   TextField "Text field_22" at 649,435 size 53x20; Text 'IW230'
   Button "HmiScreenItemData_8" at 469,45 size 355x40; TextOn 'Back'; TextOff 'Text'
   TextField "Screen title" at 455,41 size 373x50; Text 'Screen title'

screen "RIO 4 Analogue Settings" 1280x800, template "Template"
   on GenerateScreen: "TitleUpdater"()
   Button "HmiScreenItemData_1" at 1,1 size 150x40; TextOn 'Back'; TextOff 'Commissioning'
      on Release: ActivateScreen("Commissioning Main Page", 0)
   TextField "Text field_82" at 60,138 size 215x20; Text 'Tank 4P USD Flow FIT-418-4P'
   TextField "Text field_90" at 286,114 size 62x18; Text 'Reading'
   IOField "I/O field_2" at 281,138 size 75x20; FormatPattern 999; Unit  Nm³/hr
      ProcessValue <- "20_TANKS_IP_DATA_RIO_04_FIRST_TANK_USD_FLOW"
   TextField "Text field_1" at 359,114 size 68x18; Text 'Low Low'
   TextField "Text field_2" at 442,114 size 34x18; Text 'Low'
   TextField "Text field_3" at 509,114 size 37x18; Text 'High'
   TextField "Text field_4" at 561,114 size 74x18; Text 'High High'
   TextField "Text field_5" at 434,92 size 74x18; Text 'Setpoints'
   TextField "Text field_6" at 7,138 size 53x20; Text 'IW260'
   TextField "Text field_7" at 60,175 size 215x20; Text 'Tank 4P MBG Flow FIT-420-4P'
   IOField "I/O field_6" at 281,175 size 75x20; FormatPattern 999; Unit  Nm³/hr
      ProcessValue <- "20_TANKS_IP_DATA_RIO_04_FIRST_TANK_MBG_FLOW"
   TextField "Text field_8" at 7,175 size 53x20; Text 'IW262'
   TextField "Text field_9" at 60,212 size 215x20; Text 'Tank 4S USD Flow FIT-417-4S'
   IOField "I/O field_11" at 281,212 size 75x20; FormatPattern 999; Unit  Nm³/hr
      ProcessValue <- "20_TANKS_IP_DATA_RIO_04_SECOND_TANK_USD_FLOW"
   TextField "Text field_10" at 7,212 size 53x20; Text 'IW264'
   TextField "Text field_11" at 60,249 size 215x20; Text 'Tank 4S MBG Flow FIT-419-4S'
   IOField "I/O field_16" at 281,249 size 75x20; FormatPattern 999; Unit  Nm³/hr
      ProcessValue <- "20_TANKS_IP_DATA_RIO_04_SECOND_TANK_MBG_FLOW"
   TextField "Text field_12" at 7,249 size 53x20; Text 'IW266'
   TextField "Text field_13" at 60,286 size 215x20; Text 'RIO 4 Deck Main Pressure PT-415'
   TextField "Text field_14" at 7,286 size 53x20; Text 'IW268'
   TextField "Text field_15" at 60,324 size 215x20; Text 'Tank 4P BW Level LT-422-4P'
   TextField "Text field_16" at 7,324 size 53x20; Text 'IW270'
   TextField "Text field_17" at 60,361 size 215x20; Text 'Tank 4S BW Level LT-421-4S'
   TextField "Text field_18" at 7,361 size 53x20; Text 'IW272'
   TextField "Text field_25" at 702,324 size 215x20; Text 'Tank 4S BW Temperature 425-4S'
   TextField "Text field_26" at 928,114 size 62x18; Text 'Reading'
   IOField "I/O field_51" at 922,324 size 75x20; FormatPattern s999.9; Unit  °C
      ProcessValue <- "20_TANKS_IP_DATA_RIO_04_SECOND_TANK_BWT_TEMP"
   TextField "Text field_27" at 1001,114 size 68x18; Text 'Low Low'
   TextField "Text field_28" at 1082,114 size 34x18; Text 'Low'
   TextField "Text field_29" at 1150,114 size 37x18; Text 'High'
   TextField "Text field_30" at 1203,114 size 74x18; Text 'High High'
   TextField "Text field_31" at 1076,92 size 74x18; Text 'Setpoints'
   TextField "Text field_32" at 649,324 size 53x20; Text 'IW286'
   TextField "Text field_33" at 702,361 size 215x20; Text 'Tank 4S BW DO TX-427-4S'
   IOField "I/O field_56" at 922,361 size 75x20; FormatPattern 99.9; Unit  mg/l
      ProcessValue <- "20_TANKS_IP_DATA_RIO_04_SECOND_TANK_BWT_DO"
   TextField "Text field_34" at 649,361 size 53x20; Text 'IW288'
   TextField "Text field_35" at 702,398 size 215x20; Text 'Confined Space O2 Level Port'
   IOField "I/O field_61" at 922,398 size 75x20; FormatPattern 99.9; Unit  %
      ProcessValue <- "20_TANKS_IP_DATA_RIO_04_FIRST_TANK_O2_MONITOR"
   TextField "Text field_36" at 649,398 size 53x20; Text 'IW290'
   TextField "Text field_65" at 702,138 size 215x20; Text 'Tank 4P BW ph TX-426-4P'
   IOField "I/O field_126" at 922,138 size 75x20; FormatPattern 999.9
      ProcessValue <- "20_TANKS_IP_DATA_RIO_04_FIRST_TANK_BWT_PH"
   TextField "Text field_66" at 649,138 size 53x20; Text 'IW276'
   TextField "Text field_67" at 702,175 size 215x20; Text 'Tank 4P BW Temperature 426-4P'
   IOField "I/O field_131" at 922,175 size 75x20; FormatPattern s999.9; Unit  °C
      ProcessValue <- "20_TANKS_IP_DATA_RIO_04_FIRST_TANK_BWT_TEMP"
   TextField "Text field_68" at 649,175 size 53x20; Text 'IW278'
   TextField "Text field_69" at 702,212 size 215x20; Text 'Tank 4P BW DO TX-428-4P'
   IOField "I/O field_136" at 922,212 size 75x20; FormatPattern 99.9; Unit  mg/l
      ProcessValue <- "20_TANKS_IP_DATA_RIO_04_FIRST_TANK_BWT_DO"
   TextField "Text field_70" at 649,212 size 53x20; Text 'IW280'
   TextField "Text field_71" at 702,249 size 215x20; Text 'RIO 4 Tanks Pressure PT-424'
   TextField "Text field_72" at 649,249 size 53x20; Text 'IW282'
   TextField "Text field_73" at 702,286 size 215x20; Text 'Tank 4S BW ph TX-425-4S'
   IOField "I/O field_146" at 922,286 size 75x20; FormatPattern 999.9
      ProcessValue <- "20_TANKS_IP_DATA_RIO_04_SECOND_TANK_BWT_PH"
   TextField "Text field_74" at 649,286 size 53x20; Text 'IW284'
   TextField "Text field_41" at 133,114 size 85x18; Text 'Description'
   TextField "Text field_42" at 771,114 size 85x18; Text 'Description'
   TextField "Text field_43" at 17,114 size 21x18; Text 'AI'
   TextField "Text field_44" at 661,114 size 21x18; Text 'AI'
   IOField "I/O field_21" at 281,285 size 75x20; FormatPattern 99.9; Unit  Bar
      ProcessValue <- "20_TANKS_IP_DATA_RIO_04_FIRST_TANK_DECK_IG_PRESS"
   IOField "I/O field_26" at 281,322 size 75x20; FormatPattern 999.9; Unit  %
      ProcessValue <- "20_TANKS_IP_DATA_RIO_04_FIRST_TANK_BWT_LEVEL"
   IOField "I/O field_27" at 281,359 size 75x20; FormatPattern 999.9; Unit  %
      ProcessValue <- "20_TANKS_IP_DATA_RIO_04_SECOND_TANK_BWT_LEVEL"
   IOField "I/O field_93" at 922,249 size 75x20; FormatPattern s999.9; Unit  mBar
      ProcessValue <- "20_TANKS_IP_DATA_RIO_04_FIRST_TANK_TANKS_PRESS"
   TextField "Text field_21" at 702,435 size 215x20; Text 'Confined Space O2 Level Starboard'
   IOField "I/O field_41" at 922,435 size 75x20; FormatPattern 99.9; Unit  %
      ProcessValue <- "20_TANKS_IP_DATA_RIO_04_SECOND_TANK_O2_MONITOR"
   TextField "Text field_22" at 649,435 size 53x20; Text 'IW290'
   IOField "I/O field_1" at 361,138 size 60x20; Authorization "User administration"; FormatPattern 999
      ProcessValue <- "2084_Setpoints_FIT418_LoLo"
   IOField "I/O field_3" at 429,138 size 60x20; Authorization "User administration"; FormatPattern 999
      ProcessValue <- "2084_Setpoints_FIT418_Lo"
   IOField "I/O field_4" at 497,138 size 60x20; Authorization "User administration"; FormatPattern 999
      ProcessValue <- "2084_Setpoints_FIT418_Hi"
   IOField "I/O field_5" at 565,138 size 60x20; Authorization "User administration"; FormatPattern 999
      ProcessValue <- "2084_Setpoints_FIT418_HiHi"
   IOField "I/O field_7" at 361,175 size 60x20; FormatPattern 999
      ProcessValue <- "2084_Setpoints_FIT420_LoLo"
   IOField "I/O field_8" at 429,175 size 60x20; FormatPattern 999
      ProcessValue <- "2084_Setpoints_FIT420_Lo"
   IOField "I/O field_9" at 497,175 size 60x20; Authorization "User administration"; FormatPattern 999
      ProcessValue <- "2084_Setpoints_FIT420_Hi"
   IOField "I/O field_10" at 565,175 size 60x20; Authorization "User administration"; FormatPattern 999
      ProcessValue <- "2084_Setpoints_FIT420_HiHi"
   IOField "I/O field_12" at 361,212 size 60x20; FormatPattern 999
      ProcessValue <- "2084_Setpoints_FIT417_LoLo"
   IOField "I/O field_13" at 429,212 size 60x20; FormatPattern 999
      ProcessValue <- "2084_Setpoints_FIT417_Lo"
   IOField "I/O field_14" at 497,212 size 60x20; Authorization "User administration"; FormatPattern 999
      ProcessValue <- "2084_Setpoints_FIT417_Hi"
   IOField "I/O field_15" at 565,212 size 60x20; Authorization "User administration"; FormatPattern 999
      ProcessValue <- "2084_Setpoints_FIT417_HiHi"
   IOField "I/O field_17" at 361,249 size 60x20; FormatPattern 999
      ProcessValue <- "2084_Setpoints_FIT419_LoLo"
   IOField "I/O field_18" at 429,249 size 60x20; FormatPattern 999
      ProcessValue <- "2084_Setpoints_FIT419_Lo"
   IOField "I/O field_19" at 497,249 size 60x20; FormatPattern 999
      ProcessValue <- "2084_Setpoints_FIT419_Hi"
   IOField "I/O field_20" at 565,249 size 60x20; FormatPattern 999
      ProcessValue <- "2084_Setpoints_FIT419_HiHi"
   IOField "I/O field_22" at 361,285 size 60x20; FormatPattern 99.999
      ProcessValue <- "2084_Setpoints_PIT415_LoLo"
   IOField "I/O field_23" at 429,285 size 60x20; FormatPattern 99.999
      ProcessValue <- "2084_Setpoints_PIT415_Lo"
   IOField "I/O field_24" at 497,285 size 60x20; FormatPattern 99.999
      ProcessValue <- "2084_Setpoints_PIT415_Hi"
   IOField "I/O field_25" at 565,285 size 60x20; FormatPattern 99.999
      ProcessValue <- "2084_Setpoints_PIT415_HiHi"
   IOField "I/O field_28" at 429,359 size 60x20; Authorization "User administration"; FormatPattern 999
      ProcessValue <- "2084_Setpoints_LT421_Lo"
   IOField "I/O field_29" at 497,359 size 60x20; Authorization "User administration"; FormatPattern 999
      ProcessValue <- "2084_Setpoints_LT421_Hi"
   IOField "I/O field_30" at 429,322 size 60x20; Authorization "User administration"; FormatPattern 999
      ProcessValue <- "2084_Setpoints_LT422_Lo"
   IOField "I/O field_31" at 497,322 size 60x20; Authorization "User administration"; FormatPattern 999
      ProcessValue <- "2084_Setpoints_LT422_Hi"
   IOField "I/O field_32" at 361,322 size 60x20; FormatPattern 9.9
   IOField "I/O field_33" at 361,359 size 60x20; FormatPattern 9.9
   IOField "I/O field_34" at 565,322 size 60x20; FormatPattern 9.9
   IOField "I/O field_35" at 565,359 size 60x20; FormatPattern 9.9
   IOField "I/O field_62" at 1004,397 size 60x20; FormatPattern 99.9
      ProcessValue <- "2084_Setpoints_Conf O2 Level Lo Lo"
   IOField "I/O field_63" at 1072,397 size 60x20; FormatPattern 99.9
      ProcessValue <- "2084_Setpoints_Conf O2 Level Lo"
   IOField "I/O field_64" at 1139,397 size 60x20; Authorization "User administration"; FormatPattern 99.9
   IOField "I/O field_65" at 1207,397 size 60x20; Authorization "User administration"; FormatPattern 99.9
   IOField "I/O field_72" at 1004,286 size 60x20; FormatPattern 99.9
   IOField "I/O field_74" at 1004,323 size 60x20; FormatPattern 99.9
   IOField "I/O field_75" at 1072,323 size 60x20; FormatPattern 99.9
   IOField "I/O field_77" at 1207,286 size 60x20; Authorization "User administration"; FormatPattern 99.9
   IOField "I/O field_78" at 1139,323 size 60x20; Authorization "User administration"; FormatPattern 99.9
   IOField "I/O field_79" at 1207,323 size 60x20; Authorization "User administration"; FormatPattern 99.9
   IOField "I/O field_80" at 1139,360 size 60x20; Authorization "User administration"; FormatPattern 99.9
      ProcessValue <- "2084_Setpoints_TX427 Star DO High"
   IOField "I/O field_86" at 1207,360 size 60x20; Authorization "User administration"; FormatPattern 99.9
   IOField "I/O field_87" at 1004,360 size 60x20; Authorization "User administration"; FormatPattern 99.9
   IOField "I/O field_88" at 1072,360 size 60x20; Authorization "User administration"; FormatPattern 99.9
      ProcessValue <- "2084_Setpoints_TX427 Star DO Lo"
   IOField "I/O field_52" at 1003,138 size 60x20; FormatPattern 99.9
   IOField "I/O field_53" at 1071,138 size 60x20; FormatPattern 99.9
      ProcessValue <- "2084_Setpoints_TX426 Port PH Lo"
   IOField "I/O field_54" at 1003,175 size 60x20; FormatPattern 99.9
   IOField "I/O field_55" at 1071,175 size 60x20; FormatPattern 99.9
   IOField "I/O field_57" at 1139,138 size 60x20; Authorization "User administration"; FormatPattern 99.9
      ProcessValue <- "2084_Setpoints_TX426 Port PH High"
   IOField "I/O field_58" at 1207,138 size 60x20; Authorization "User administration"; FormatPattern 99.9
   IOField "I/O field_59" at 1139,175 size 60x20; Authorization "User administration"; FormatPattern 99.9
   IOField "I/O field_60" at 1207,175 size 60x20; Authorization "User administration"; FormatPattern 99.9
   IOField "I/O field_89" at 1139,212 size 60x20; Authorization "User administration"; FormatPattern 99.9
      ProcessValue <- "2084_Setpoints_TX428 Port DO High"
   IOField "I/O field_90" at 1207,212 size 60x20; Authorization "User administration"; FormatPattern 99.9
   IOField "I/O field_91" at 1003,212 size 60x20; Authorization "User administration"; FormatPattern 99.9
   IOField "I/O field_92" at 1071,212 size 60x20; Authorization "User administration"; FormatPattern 99.9
      ProcessValue <- "2084_Setpoints_TX428 Port DO Lo"
   IOField "I/O field_94" at 1139,249 size 60x20; Authorization "User administration"; FormatPattern 999.9
      ProcessValue <- "2084_Setpoints_PIT424_Hi"
   IOField "I/O field_95" at 1207,249 size 60x20; Authorization "User administration"; FormatPattern 999.9
      ProcessValue <- "2084_Setpoints_PIT424_HiHi"
   IOField "I/O field_96" at 1004,249 size 60x20; Authorization "User administration"; FormatPattern 999.9
      ProcessValue <- "2084_Setpoints_PIT424_LoLo"
   IOField "I/O field_97" at 1072,249 size 60x20; Authorization "User administration"; FormatPattern 999.9
      ProcessValue <- "2084_Setpoints_PIT424_Lo"
   IOField "I/O field_42" at 1072,286 size 60x20; FormatPattern 99.9
      ProcessValue <- "2084_Setpoints_TX425 Star PH Lo"
   IOField "I/O field_43" at 1139,286 size 60x20; Authorization "User administration"; FormatPattern 99.9
      ProcessValue <- "2084_Setpoints_TX425 Star PH High"
   Group "Group" at 455,41 size 373x50
   Button "HmiScreenItemData_8" at 469,45 size 355x40; TextOn 'Back'; TextOff 'Text'
   TextField "Screen title" at 455,41 size 373x50; Text 'Screen title'

screen "RIO 5 Analogue Settings" 1280x800, template "Template"
   on GenerateScreen: "TitleUpdater"()
   Button "HmiScreenItemData_1" at 1,1 size 150x40; TextOn 'Back'; TextOff 'Commissioning'
      on Release: ActivateScreen("Commissioning Main Page", 0)
   TextField "Text field_82" at 60,138 size 215x20; Text 'Tank 5P USD Flow FIT-418-5P'
   TextField "Text field_90" at 286,114 size 62x18; Text 'Reading'
   IOField "I/O field_2" at 281,138 size 75x20; FormatPattern 999; Unit  Nm³/hr
      ProcessValue <- "20_TANKS_IP_DATA_RIO_05_FIRST_TANK_USD_FLOW"
   TextField "Text field_1" at 359,114 size 68x18; Text 'Low Low'
   TextField "Text field_2" at 442,114 size 34x18; Text 'Low'
   TextField "Text field_3" at 509,114 size 37x18; Text 'High'
   TextField "Text field_4" at 561,114 size 74x18; Text 'High High'
   TextField "Text field_5" at 434,92 size 74x18; Text 'Setpoints'
   TextField "Text field_6" at 7,138 size 53x20; Text 'IW300'
   TextField "Text field_7" at 60,175 size 215x20; Text 'Tank 5P MBG Flow FIT-420-5P'
   IOField "I/O field_6" at 281,175 size 75x20; FormatPattern 999; Unit  Nm³/hr
      ProcessValue <- "20_TANKS_IP_DATA_RIO_05_FIRST_TANK_MBG_FLOW"
   TextField "Text field_8" at 7,175 size 53x20; Text 'IW302'
   TextField "Text field_9" at 60,212 size 215x20; Text 'Tank 5S USD Flow FIT-417-5S'
   IOField "I/O field_11" at 281,212 size 75x20; FormatPattern 999; Unit  Nm³/hr
      ProcessValue <- "20_TANKS_IP_DATA_RIO_05_SECOND_TANK_USD_FLOW"
   TextField "Text field_10" at 7,212 size 53x20; Text 'IW304'
   TextField "Text field_11" at 60,249 size 215x20; Text 'Tank 5S MBG Flow FIT-419-5S'
   IOField "I/O field_16" at 281,249 size 75x20; FormatPattern 999; Unit  Nm³/hr
      ProcessValue <- "20_TANKS_IP_DATA_RIO_05_SECOND_TANK_MBG_FLOW"
   TextField "Text field_12" at 7,249 size 53x20; Text 'IW306'
   TextField "Text field_13" at 60,286 size 215x20; Text 'RIO 5 Deck Main Pressure PT-415'
   TextField "Text field_14" at 7,286 size 53x20; Text 'IW308'
   TextField "Text field_15" at 60,324 size 215x20; Text 'Tank 5P BW Level LT-422-5P'
   TextField "Text field_16" at 7,324 size 53x20; Text 'IW310'
   TextField "Text field_17" at 60,361 size 215x20; Text 'Tank 5S BW Level LT-421-5S'
   TextField "Text field_18" at 7,361 size 53x20; Text 'IW312'
   TextField "Text field_25" at 702,324 size 215x20; Text 'Tank 5S BW Temperature 425-5S'
   TextField "Text field_26" at 928,114 size 62x18; Text 'Reading'
   IOField "I/O field_51" at 922,324 size 75x20; FormatPattern s999.9; Unit  °C
      ProcessValue <- "20_TANKS_IP_DATA_RIO_05_SECOND_TANK_BWT_TEMP"
   TextField "Text field_27" at 1001,114 size 68x18; Text 'Low Low'
   TextField "Text field_28" at 1082,114 size 34x18; Text 'Low'
   TextField "Text field_29" at 1150,114 size 37x18; Text 'High'
   TextField "Text field_30" at 1203,114 size 74x18; Text 'High High'
   TextField "Text field_31" at 1076,92 size 74x18; Text 'Setpoints'
   TextField "Text field_32" at 649,324 size 53x20; Text 'IW326'
   TextField "Text field_33" at 702,361 size 215x20; Text 'Tank 5S BW DO TX-427-5S'
   IOField "I/O field_56" at 922,361 size 75x20; FormatPattern 99.9; Unit  mg/l
      ProcessValue <- "20_TANKS_IP_DATA_RIO_05_SECOND_TANK_BWT_DO"
   TextField "Text field_34" at 649,361 size 53x20; Text 'IW328'
   TextField "Text field_35" at 702,398 size 215x20; Text 'Confined Space Oxygen Level'
   IOField "I/O field_61" at 922,398 size 75x20; FormatPattern 99.9; Unit  %
      ProcessValue <- "20_TANKS_IP_DATA_RIO_05_FIRST_TANK_O2_MONITOR"
   TextField "Text field_36" at 649,398 size 53x20; Text 'IW330'
   TextField "Text field_65" at 702,138 size 215x20; Text 'Tank 5P BW ph TX-426-5P'
   IOField "I/O field_126" at 922,138 size 75x20; FormatPattern 99.9
      ProcessValue <- "20_TANKS_IP_DATA_RIO_05_FIRST_TANK_BWT_PH"
   TextField "Text field_66" at 649,138 size 53x20; Text 'IW316'
   TextField "Text field_67" at 702,175 size 215x20; Text 'Tank 5P BW Temperature 426-5P'
   IOField "I/O field_131" at 922,175 size 75x20; FormatPattern s999.9; Unit  °C
      ProcessValue <- "20_TANKS_IP_DATA_RIO_05_FIRST_TANK_BWT_TEMP"
   TextField "Text field_68" at 649,175 size 53x20; Text 'IW318'
   TextField "Text field_69" at 702,212 size 215x20; Text 'Tank 5P BW DO TX-428-5P'
   IOField "I/O field_136" at 922,212 size 75x20; FormatPattern s99.99; Unit  mg/l
      ProcessValue <- "20_TANKS_IP_DATA_RIO_05_FIRST_TANK_BWT_DO"
   TextField "Text field_70" at 649,212 size 53x20; Text 'IW320'
   TextField "Text field_71" at 702,249 size 215x20; Text 'RIO 5 Tanks Pressure PT-424'
   TextField "Text field_72" at 649,249 size 53x20; Text 'IW322'
   TextField "Text field_73" at 702,286 size 215x20; Text 'Tank 5S BW ph TX-425-5S'
   IOField "I/O field_146" at 922,286 size 75x20; FormatPattern 99.9
      ProcessValue <- "20_TANKS_IP_DATA_RIO_05_SECOND_TANK_BWT_PH"
   TextField "Text field_74" at 649,286 size 53x20; Text 'IW324'
   TextField "Text field_41" at 133,114 size 85x18; Text 'Description'
   TextField "Text field_42" at 771,114 size 85x18; Text 'Description'
   TextField "Text field_43" at 17,114 size 21x18; Text 'AI'
   TextField "Text field_44" at 661,114 size 21x18; Text 'AI'
   IOField "I/O field_21" at 281,285 size 75x20; FormatPattern 99.999; Unit  Bar
      ProcessValue <- "20_TANKS_IP_DATA_RIO_05_FIRST_TANK_DECK_IG_PRESS"
   IOField "I/O field_26" at 281,322 size 75x20; FormatPattern 999.9; Unit  %
      ProcessValue <- "20_TANKS_IP_DATA_RIO_05_FIRST_TANK_BWT_LEVEL"
   IOField "I/O field_27" at 281,359 size 75x20; FormatPattern 999.9; Unit  %
      ProcessValue <- "20_TANKS_IP_DATA_RIO_05_SECOND_TANK_BWT_LEVEL"
   IOField "I/O field_93" at 922,249 size 75x20; FormatPattern 999.9; Unit  mBar
      ProcessValue <- "20_TANKS_IP_DATA_RIO_05_FIRST_TANK_TANKS_PRESS"
   Group "Group" at 455,41 size 373x50
   TextField "Text field_21" at 702,435 size 215x20; Text 'Confined Space Oxygen Level'
   IOField "I/O field_41" at 922,435 size 75x20; FormatPattern 99.9; Unit  %
      ProcessValue <- "20_TANKS_IP_DATA_RIO_05_SECOND_TANK_O2_MONITOR"
   TextField "Text field_22" at 649,435 size 53x20; Text 'IW330'
   IOField "I/O field_1" at 361,138 size 60x20; Authorization "User administration"; FormatPattern 999
      ProcessValue <- "2084_Setpoints_FIT418_LoLo"
   IOField "I/O field_3" at 429,138 size 60x20; Authorization "User administration"; FormatPattern 999
      ProcessValue <- "2084_Setpoints_FIT418_Lo"
   IOField "I/O field_4" at 497,138 size 60x20; Authorization "User administration"; FormatPattern 999
      ProcessValue <- "2084_Setpoints_FIT418_Hi"
   IOField "I/O field_5" at 565,138 size 60x20; Authorization "User administration"; FormatPattern 999
      ProcessValue <- "2084_Setpoints_FIT418_HiHi"
   IOField "I/O field_7" at 361,175 size 60x20; FormatPattern 999
      ProcessValue <- "2084_Setpoints_FIT420_LoLo"
   IOField "I/O field_8" at 429,175 size 60x20; FormatPattern 999
      ProcessValue <- "2084_Setpoints_FIT420_Lo"
   IOField "I/O field_9" at 497,175 size 60x20; Authorization "User administration"; FormatPattern 999
      ProcessValue <- "2084_Setpoints_FIT420_Hi"
   IOField "I/O field_10" at 565,175 size 60x20; Authorization "User administration"; FormatPattern 999
      ProcessValue <- "2084_Setpoints_FIT420_HiHi"
   IOField "I/O field_12" at 361,212 size 60x20; FormatPattern 999
      ProcessValue <- "2084_Setpoints_FIT417_LoLo"
   IOField "I/O field_13" at 429,212 size 60x20; FormatPattern 999
      ProcessValue <- "2084_Setpoints_FIT417_Lo"
   IOField "I/O field_14" at 497,212 size 60x20; Authorization "User administration"; FormatPattern 999
      ProcessValue <- "2084_Setpoints_FIT417_Hi"
   IOField "I/O field_15" at 565,212 size 60x20; Authorization "User administration"; FormatPattern 999
      ProcessValue <- "2084_Setpoints_FIT417_HiHi"
   IOField "I/O field_17" at 361,249 size 60x20; FormatPattern 999
      ProcessValue <- "2084_Setpoints_FIT419_LoLo"
   IOField "I/O field_18" at 429,249 size 60x20; FormatPattern 999
      ProcessValue <- "2084_Setpoints_FIT419_Lo"
   IOField "I/O field_19" at 497,249 size 60x20; FormatPattern 999
      ProcessValue <- "2084_Setpoints_FIT419_Hi"
   IOField "I/O field_20" at 565,249 size 60x20; FormatPattern 999
      ProcessValue <- "2084_Setpoints_FIT419_HiHi"
   IOField "I/O field_22" at 361,285 size 60x20; FormatPattern 99.999
      ProcessValue <- "2084_Setpoints_PIT415_LoLo"
   IOField "I/O field_23" at 429,285 size 60x20; FormatPattern 99.999
      ProcessValue <- "2084_Setpoints_PIT415_Lo"
   IOField "I/O field_24" at 497,285 size 60x20; FormatPattern 99.999
      ProcessValue <- "2084_Setpoints_PIT415_Hi"
   IOField "I/O field_25" at 565,285 size 60x20; FormatPattern 99.999
      ProcessValue <- "2084_Setpoints_PIT415_HiHi"
   IOField "I/O field_28" at 429,359 size 60x20; Authorization "User administration"; FormatPattern 999
      ProcessValue <- "2084_Setpoints_LT421_Lo"
   IOField "I/O field_29" at 497,359 size 60x20; Authorization "User administration"; FormatPattern 999
      ProcessValue <- "2084_Setpoints_LT421_Hi"
   IOField "I/O field_30" at 429,322 size 60x20; Authorization "User administration"; FormatPattern 999
      ProcessValue <- "2084_Setpoints_LT422_Lo"
   IOField "I/O field_31" at 497,322 size 60x20; Authorization "User administration"; FormatPattern 999
      ProcessValue <- "2084_Setpoints_LT422_Hi"
   IOField "I/O field_32" at 361,322 size 60x20; FormatPattern 9.9
   IOField "I/O field_33" at 361,359 size 60x20; FormatPattern 9.9
   IOField "I/O field_34" at 565,322 size 60x20; FormatPattern 9.9
   IOField "I/O field_35" at 565,359 size 60x20; FormatPattern 9.9
   IOField "I/O field_62" at 1004,397 size 60x20; FormatPattern 99.9
      ProcessValue <- "2084_Setpoints_Conf O2 Level Lo Lo"
   IOField "I/O field_63" at 1072,397 size 60x20; FormatPattern 99.9
      ProcessValue <- "2084_Setpoints_Conf O2 Level Lo"
   IOField "I/O field_64" at 1139,397 size 60x20; Authorization "User administration"; FormatPattern 99.9
   IOField "I/O field_65" at 1207,397 size 60x20; Authorization "User administration"; FormatPattern 99.9
   IOField "I/O field_72" at 1004,286 size 60x20; FormatPattern 99.9
   IOField "I/O field_74" at 1004,323 size 60x20; FormatPattern 99.9
   IOField "I/O field_75" at 1072,323 size 60x20; FormatPattern 99.9
   IOField "I/O field_77" at 1207,286 size 60x20; Authorization "User administration"; FormatPattern 99.9
   IOField "I/O field_78" at 1139,323 size 60x20; Authorization "User administration"; FormatPattern 99.9
   IOField "I/O field_79" at 1207,323 size 60x20; Authorization "User administration"; FormatPattern 99.9
   IOField "I/O field_80" at 1139,360 size 60x20; Authorization "User administration"; FormatPattern 99.9
      ProcessValue <- "2084_Setpoints_TX427 Star DO High"
   IOField "I/O field_86" at 1207,360 size 60x20; Authorization "User administration"; FormatPattern 99.9
   IOField "I/O field_87" at 1004,360 size 60x20; Authorization "User administration"; FormatPattern 99.9
   IOField "I/O field_88" at 1072,360 size 60x20; Authorization "User administration"; FormatPattern 99.9
      ProcessValue <- "2084_Setpoints_TX427 Star DO Lo"
   IOField "I/O field_52" at 1003,138 size 60x20; FormatPattern 99.9
   IOField "I/O field_53" at 1071,138 size 60x20; FormatPattern 99.9
      ProcessValue <- "2084_Setpoints_TX426 Port PH Lo"
   IOField "I/O field_54" at 1003,175 size 60x20; FormatPattern 99.9
   IOField "I/O field_55" at 1071,175 size 60x20; FormatPattern 99.9
   IOField "I/O field_57" at 1139,138 size 60x20; Authorization "User administration"; FormatPattern 99.9
      ProcessValue <- "2084_Setpoints_TX426 Port PH High"
   IOField "I/O field_58" at 1207,138 size 60x20; Authorization "User administration"; FormatPattern 99.9
   IOField "I/O field_59" at 1139,175 size 60x20; Authorization "User administration"; FormatPattern 99.9
   IOField "I/O field_60" at 1207,175 size 60x20; Authorization "User administration"; FormatPattern 99.9
   IOField "I/O field_89" at 1139,212 size 60x20; Authorization "User administration"; FormatPattern 99.9
      ProcessValue <- "2084_Setpoints_TX428 Port DO High"
   IOField "I/O field_90" at 1207,212 size 60x20; Authorization "User administration"; FormatPattern 99.9
   IOField "I/O field_91" at 1003,212 size 60x20; Authorization "User administration"; FormatPattern 99.9
   IOField "I/O field_92" at 1071,212 size 60x20; Authorization "User administration"; FormatPattern 99.9
      ProcessValue <- "2084_Setpoints_TX428 Port DO Lo"
   IOField "I/O field_94" at 1139,249 size 60x20; Authorization "User administration"; FormatPattern 999.9
      ProcessValue <- "2084_Setpoints_PIT424_Hi"
   IOField "I/O field_95" at 1207,249 size 60x20; Authorization "User administration"; FormatPattern 999.9
      ProcessValue <- "2084_Setpoints_PIT424_HiHi"
   IOField "I/O field_96" at 1004,249 size 60x20; Authorization "User administration"; FormatPattern 999.9
      ProcessValue <- "2084_Setpoints_PIT424_LoLo"
   IOField "I/O field_97" at 1072,249 size 60x20; Authorization "User administration"; FormatPattern 999.9
      ProcessValue <- "2084_Setpoints_PIT424_Lo"
   IOField "I/O field_36" at 1072,286 size 60x20; FormatPattern 99.9
      ProcessValue <- "2084_Setpoints_TX425 Star PH Lo"
   IOField "I/O field_42" at 1139,286 size 60x20; Authorization "User administration"; FormatPattern 99.9
      ProcessValue <- "2084_Setpoints_TX425 Star PH High"
   Button "HmiScreenItemData_8" at 469,45 size 355x40; TextOn 'Back'; TextOff 'Text'
   TextField "Screen title" at 455,41 size 373x50; Text 'Screen title'

screen "RIO 6 Analogue Settings" 1280x800, template "Template"
   on GenerateScreen: "TitleUpdater"()
   Button "HmiScreenItemData_1" at 1,1 size 150x40; TextOn 'Back'; TextOff 'Commissioning'
      on Release: ActivateScreen("Commissioning Main Page", 0)
   TextField "Text field_82" at 60,138 size 215x20; Text 'Tank 6P USD Flow FIT-418-6P'
   TextField "Text field_90" at 286,114 size 62x18; Text 'Reading'
   IOField "I/O field_2" at 281,138 size 75x20; FormatPattern 999; Unit  Nm³/hr
      ProcessValue <- "20_TANKS_IP_DATA_RIO_06_FIRST_TANK_USD_FLOW"
   TextField "Text field_1" at 359,114 size 68x18; Text 'Low Low'
   TextField "Text field_2" at 442,114 size 34x18; Text 'Low'
   TextField "Text field_3" at 509,114 size 37x18; Text 'High'
   TextField "Text field_4" at 561,114 size 74x18; Text 'High High'
   TextField "Text field_5" at 434,92 size 74x18; Text 'Setpoints'
   TextField "Text field_6" at 7,138 size 53x20; Text 'IW360'
   TextField "Text field_7" at 60,175 size 215x20; Text 'Tank 6P MBG Flow FIT-420-6P'
   IOField "I/O field_6" at 281,175 size 75x20; FormatPattern 999; Unit  Nm³/hr
      ProcessValue <- "20_TANKS_IP_DATA_RIO_06_FIRST_TANK_MBG_FLOW"
   TextField "Text field_8" at 7,175 size 53x20; Text 'IW362'
   TextField "Text field_9" at 60,212 size 215x20; Text 'Tank 6S USD Flow FIT-417-6S'
   IOField "I/O field_11" at 281,212 size 75x20; FormatPattern 999; Unit  Nm³/hr
      ProcessValue <- "20_TANKS_IP_DATA_RIO_06_SECOND_TANK_USD_FLOW"
   TextField "Text field_10" at 7,212 size 53x20; Text 'IW364'
   TextField "Text field_11" at 60,249 size 215x20; Text 'Tank 6S MBG Flow FIT-419-6S'
   IOField "I/O field_16" at 281,249 size 75x20; FormatPattern 999; Unit  Nm³/hr
      ProcessValue <- "20_TANKS_IP_DATA_RIO_06_SECOND_TANK_MBG_FLOW"
   TextField "Text field_12" at 7,249 size 53x20; Text 'IW366'
   TextField "Text field_13" at 60,286 size 215x20; Text 'RIO 6 Deck Main Pressure PT-415'
   TextField "Text field_14" at 7,286 size 53x20; Text 'IW368'
   TextField "Text field_15" at 60,324 size 215x20; Text 'Tank 6P BW Level LT-422-6P'
   TextField "Text field_16" at 7,324 size 53x20; Text 'IW370'
   TextField "Text field_17" at 60,361 size 215x20; Text 'Tank 6S BW Level LT-421-6S'
   TextField "Text field_18" at 7,361 size 53x20; Text 'IW372'
   TextField "Text field_25" at 702,324 size 215x20; Text 'Tank 6S BW Temperature 425-6S'
   TextField "Text field_26" at 928,114 size 62x18; Text 'Reading'
   IOField "I/O field_51" at 922,324 size 75x20; FormatPattern s999.9; Unit  °C
      ProcessValue <- "20_TANKS_IP_DATA_RIO_06_SECOND_TANK_BWT_TEMP"
   TextField "Text field_27" at 1001,114 size 68x18; Text 'Low Low'
   TextField "Text field_28" at 1082,114 size 34x18; Text 'Low'
   TextField "Text field_29" at 1150,114 size 37x18; Text 'High'
   TextField "Text field_30" at 1203,114 size 74x18; Text 'High High'
   TextField "Text field_31" at 1076,92 size 74x18; Text 'Setpoints'
   TextField "Text field_32" at 649,324 size 53x20; Text 'IW386'
   TextField "Text field_33" at 702,361 size 215x20; Text 'Tank 6S BW DO TX-427-6S'
   IOField "I/O field_56" at 922,361 size 75x20; FormatPattern 99.9; Unit  mg/l
      ProcessValue <- "20_TANKS_IP_DATA_RIO_06_SECOND_TANK_BWT_DO"
   TextField "Text field_34" at 649,361 size 53x20; Text 'IW388'
   TextField "Text field_35" at 702,398 size 215x20; Text 'Confined Space Oxygen Level'
   IOField "I/O field_61" at 922,398 size 75x20; FormatPattern 99.9; Unit  %
      ProcessValue <- "20_TANKS_IP_DATA_RIO_06_FIRST_TANK_O2_MONITOR"
   TextField "Text field_36" at 649,398 size 53x20; Text 'IW390'
   TextField "Text field_65" at 702,138 size 215x20; Text 'Tank 6P BW ph TX-426-6P'
   IOField "I/O field_126" at 922,138 size 75x20; FormatPattern 99.9
      ProcessValue <- "20_TANKS_IP_DATA_RIO_06_FIRST_TANK_BWT_PH"
   TextField "Text field_66" at 649,138 size 53x20; Text 'IW376'
   TextField "Text field_67" at 702,175 size 215x20; Text 'Tank 6P BW Temperature 426-6P'
   IOField "I/O field_131" at 922,175 size 75x20; FormatPattern s999.9; Unit  °C
      ProcessValue <- "20_TANKS_IP_DATA_RIO_06_FIRST_TANK_BWT_TEMP"
   TextField "Text field_68" at 649,175 size 53x20; Text 'IW378'
   TextField "Text field_69" at 702,212 size 215x20; Text 'Tank 6P BW DO TX-428-6P'
   IOField "I/O field_136" at 922,212 size 75x20; FormatPattern 99.9; Unit  mg/l
      ProcessValue <- "20_TANKS_IP_DATA_RIO_06_FIRST_TANK_BWT_DO"
   TextField "Text field_70" at 649,212 size 53x20; Text 'IW380'
   TextField "Text field_71" at 702,249 size 215x20; Text 'RIO 6 Tanks Pressure PT-424'
   TextField "Text field_72" at 649,249 size 53x20; Text 'IW382'
   TextField "Text field_73" at 702,286 size 215x20; Text 'Tank 6S BW ph TX-425-6S'
   IOField "I/O field_146" at 922,286 size 75x20; FormatPattern 99.9
      ProcessValue <- "20_TANKS_IP_DATA_RIO_06_SECOND_TANK_BWT_PH"
   TextField "Text field_74" at 649,286 size 53x20; Text 'IW384'
   TextField "Text field_41" at 133,114 size 85x18; Text 'Description'
   TextField "Text field_42" at 771,114 size 85x18; Text 'Description'
   TextField "Text field_43" at 17,114 size 21x18; Text 'AI'
   TextField "Text field_44" at 661,114 size 21x18; Text 'AI'
   IOField "I/O field_21" at 281,285 size 75x20; FormatPattern s99.999; Unit  Bar
      ProcessValue <- "20_TANKS_IP_DATA_RIO_06_FIRST_TANK_DECK_IG_PRESS"
   IOField "I/O field_26" at 281,322 size 75x20; FormatPattern 999; Unit  %
      ProcessValue <- "20_TANKS_IP_DATA_RIO_06_FIRST_TANK_BWT_LEVEL"
   IOField "I/O field_27" at 281,359 size 75x20; FormatPattern 999; Unit  %
      ProcessValue <- "20_TANKS_IP_DATA_RIO_06_SECOND_TANK_BWT_LEVEL"
   IOField "I/O field_93" at 922,249 size 75x20; FormatPattern s999.9; Unit  mBar
      ProcessValue <- "20_TANKS_IP_DATA_RIO_06_FIRST_TANK_TANKS_PRESS"
   TextField "Text field_19" at 702,434 size 215x20; Text 'Confined Space Oxygen Level'
   IOField "I/O field_36" at 922,434 size 75x20; FormatPattern 99.9; Unit  %
      ProcessValue <- "20_TANKS_IP_DATA_RIO_06_FIRST_TANK_O2_MONITOR"
   TextField "Text field_20" at 649,434 size 53x20; Text 'IW390'
   IOField "I/O field_1" at 361,138 size 60x20; Authorization "User administration"; FormatPattern 999
      ProcessValue <- "2084_Setpoints_FIT418_LoLo"
   IOField "I/O field_3" at 429,138 size 60x20; Authorization "User administration"; FormatPattern 999
      ProcessValue <- "2084_Setpoints_FIT418_Lo"
   IOField "I/O field_4" at 497,138 size 60x20; Authorization "User administration"; FormatPattern 999
      ProcessValue <- "2084_Setpoints_FIT418_Hi"
   IOField "I/O field_5" at 565,138 size 60x20; Authorization "User administration"; FormatPattern 999
      ProcessValue <- "2084_Setpoints_FIT418_HiHi"
   IOField "I/O field_7" at 361,175 size 60x20; FormatPattern 999
      ProcessValue <- "2084_Setpoints_FIT420_LoLo"
   IOField "I/O field_8" at 429,175 size 60x20; FormatPattern 999
      ProcessValue <- "2084_Setpoints_FIT420_Lo"
   IOField "I/O field_9" at 497,175 size 60x20; Authorization "User administration"; FormatPattern 999
      ProcessValue <- "2084_Setpoints_FIT420_Hi"
   IOField "I/O field_10" at 565,175 size 60x20; Authorization "User administration"; FormatPattern 999
      ProcessValue <- "2084_Setpoints_FIT420_HiHi"
   IOField "I/O field_12" at 361,212 size 60x20; FormatPattern 999
      ProcessValue <- "2084_Setpoints_FIT417_LoLo"
   IOField "I/O field_13" at 429,212 size 60x20; FormatPattern 999
      ProcessValue <- "2084_Setpoints_FIT417_Lo"
   IOField "I/O field_14" at 497,212 size 60x20; Authorization "User administration"; FormatPattern 999
      ProcessValue <- "2084_Setpoints_FIT417_Hi"
   IOField "I/O field_15" at 565,212 size 60x20; Authorization "User administration"; FormatPattern 999
      ProcessValue <- "2084_Setpoints_FIT417_HiHi"
   IOField "I/O field_17" at 361,249 size 60x20; FormatPattern 999
      ProcessValue <- "2084_Setpoints_FIT419_LoLo"
   IOField "I/O field_18" at 429,249 size 60x20; FormatPattern 999
      ProcessValue <- "2084_Setpoints_FIT419_Lo"
   IOField "I/O field_19" at 497,249 size 60x20; FormatPattern 999
      ProcessValue <- "2084_Setpoints_FIT419_Hi"
   IOField "I/O field_20" at 565,249 size 60x20; FormatPattern 999
      ProcessValue <- "2084_Setpoints_FIT419_HiHi"
   IOField "I/O field_22" at 361,285 size 60x20; FormatPattern 99.999
      ProcessValue <- "2084_Setpoints_PIT415_LoLo"
   IOField "I/O field_23" at 429,285 size 60x20; FormatPattern 99.999
      ProcessValue <- "2084_Setpoints_PIT415_Lo"
   IOField "I/O field_24" at 497,285 size 60x20; FormatPattern 99.999
      ProcessValue <- "2084_Setpoints_PIT415_Hi"
   IOField "I/O field_25" at 565,285 size 60x20; FormatPattern 99.999
      ProcessValue <- "2084_Setpoints_PIT415_HiHi"
   IOField "I/O field_28" at 429,359 size 60x20; Authorization "User administration"; FormatPattern 999
      ProcessValue <- "2084_Setpoints_LT421_Lo"
   IOField "I/O field_29" at 497,359 size 60x20; Authorization "User administration"; FormatPattern 999
      ProcessValue <- "2084_Setpoints_LT421_Hi"
   IOField "I/O field_30" at 429,322 size 60x20; Authorization "User administration"; FormatPattern 999
      ProcessValue <- "2084_Setpoints_LT422_Lo"
   IOField "I/O field_31" at 497,322 size 60x20; Authorization "User administration"; FormatPattern 999
      ProcessValue <- "2084_Setpoints_LT422_Hi"
   IOField "I/O field_32" at 361,322 size 60x20; FormatPattern 9.9
   IOField "I/O field_33" at 361,359 size 60x20; FormatPattern 9.9
   IOField "I/O field_34" at 565,322 size 60x20; FormatPattern 9.9
   IOField "I/O field_35" at 565,359 size 60x20; FormatPattern 9.9
   IOField "I/O field_62" at 1004,397 size 60x20; FormatPattern 99.9
      ProcessValue <- "2084_Setpoints_Conf O2 Level Lo Lo"
   IOField "I/O field_63" at 1072,397 size 60x20; FormatPattern 99.9
      ProcessValue <- "2084_Setpoints_Conf O2 Level Lo"
   IOField "I/O field_64" at 1139,397 size 60x20; Authorization "User administration"; FormatPattern 99.9
   IOField "I/O field_65" at 1207,397 size 60x20; Authorization "User administration"; FormatPattern 99.9
   IOField "I/O field_72" at 1004,286 size 60x20; FormatPattern 99.9
   IOField "I/O field_74" at 1004,323 size 60x20; FormatPattern 99.9
   IOField "I/O field_75" at 1072,323 size 60x20; FormatPattern 99.9
   IOField "I/O field_77" at 1207,286 size 60x20; Authorization "User administration"; FormatPattern 99.9
   IOField "I/O field_78" at 1139,323 size 60x20; Authorization "User administration"; FormatPattern 99.9
   IOField "I/O field_79" at 1207,323 size 60x20; Authorization "User administration"; FormatPattern 99.9
   IOField "I/O field_80" at 1139,360 size 60x20; Authorization "User administration"; FormatPattern 99.9
      ProcessValue <- "2084_Setpoints_TX427 Star DO High"
   IOField "I/O field_86" at 1207,360 size 60x20; Authorization "User administration"; FormatPattern 99.9
   IOField "I/O field_87" at 1004,360 size 60x20; Authorization "User administration"; FormatPattern 99.9
   IOField "I/O field_88" at 1072,360 size 60x20; Authorization "User administration"; FormatPattern 99.9
      ProcessValue <- "2084_Setpoints_TX427 Star DO Lo"
   IOField "I/O field_52" at 1003,138 size 60x20; FormatPattern 99.9
   IOField "I/O field_53" at 1071,138 size 60x20; FormatPattern 99.9
      ProcessValue <- "2084_Setpoints_TX426 Port PH Lo"
   IOField "I/O field_54" at 1003,175 size 60x20; FormatPattern 99.9
   IOField "I/O field_55" at 1071,175 size 60x20; FormatPattern 99.9
   IOField "I/O field_57" at 1139,138 size 60x20; Authorization "User administration"; FormatPattern 99.9
      ProcessValue <- "2084_Setpoints_TX426 Port PH High"
   IOField "I/O field_58" at 1207,138 size 60x20; Authorization "User administration"; FormatPattern 99.9
   IOField "I/O field_59" at 1139,175 size 60x20; Authorization "User administration"; FormatPattern 99.9
   IOField "I/O field_60" at 1207,175 size 60x20; Authorization "User administration"; FormatPattern 99.9
   IOField "I/O field_89" at 1139,212 size 60x20; Authorization "User administration"; FormatPattern 99.9
      ProcessValue <- "2084_Setpoints_TX428 Port DO High"
   IOField "I/O field_90" at 1207,212 size 60x20; Authorization "User administration"; FormatPattern 99.9
   IOField "I/O field_91" at 1003,212 size 60x20; Authorization "User administration"; FormatPattern 99.9
   IOField "I/O field_92" at 1071,212 size 60x20; Authorization "User administration"; FormatPattern 99.9
      ProcessValue <- "2084_Setpoints_TX428 Port DO Lo"
   IOField "I/O field_94" at 1139,249 size 60x20; Authorization "User administration"; FormatPattern 999.9
      ProcessValue <- "2084_Setpoints_PIT424_Hi"
   IOField "I/O field_95" at 1207,249 size 60x20; Authorization "User administration"; FormatPattern 999.9
      ProcessValue <- "2084_Setpoints_PIT424_HiHi"
   IOField "I/O field_96" at 1004,249 size 60x20; Authorization "User administration"; FormatPattern 999.9
      ProcessValue <- "2084_Setpoints_PIT424_LoLo"
   IOField "I/O field_97" at 1072,249 size 60x20; Authorization "User administration"; FormatPattern 999.9
      ProcessValue <- "2084_Setpoints_PIT424_Lo"
   IOField "I/O field_41" at 1072,286 size 60x20; FormatPattern 99.9
      ProcessValue <- "2084_Setpoints_TX425 Star PH Lo"
   IOField "I/O field_42" at 1139,286 size 60x20; Authorization "User administration"; FormatPattern 99.9
      ProcessValue <- "2084_Setpoints_TX425 Star PH High"
   Group "Group" at 455,41 size 373x50
   Button "HmiScreenItemData_8" at 469,45 size 355x40; TextOn 'Back'; TextOff 'Text'
   TextField "Screen title" at 455,41 size 373x50; Text 'Screen title'

screen "RIO 7 Analogue Settings" 1280x800, template "Template"
   on GenerateScreen: "TitleUpdater"()
   Button "HmiScreenItemData_1" at 1,1 size 150x40; TextOn 'Back'; TextOff 'Commissioning'
      on Release: ActivateScreen("Commissioning Main Page", 0)
   TextField "Text field_82" at 60,138 size 215x20; Text 'APT USD Flow FIT-418-APT'
   TextField "Text field_90" at 286,114 size 62x18; Text 'Reading'
   IOField "I/O field_2" at 281,138 size 75x20; FormatPattern 999; Unit  Nm³/hr
      ProcessValue <- "20_TANKS_IP_DATA_RIO_07_FIRST_TANK_USD_FLOW"
   TextField "Text field_1" at 359,114 size 68x18; Text 'Low Low'
   TextField "Text field_2" at 442,114 size 34x18; Text 'Low'
   TextField "Text field_3" at 509,114 size 37x18; Text 'High'
   TextField "Text field_4" at 561,114 size 74x18; Text 'High High'
   TextField "Text field_5" at 434,92 size 74x18; Text 'Setpoints'
   TextField "Text field_6" at 7,138 size 53x20; Text 'IW400'
   TextField "Text field_7" at 60,175 size 215x20; Text 'APT MBG Flow FIT-420-APT'
   IOField "I/O field_6" at 281,175 size 75x20; FormatPattern 999; Unit  Nm³/hr
      ProcessValue <- "20_TANKS_IP_DATA_RIO_07_FIRST_TANK_MBG_FLOW"
   TextField "Text field_8" at 7,175 size 53x20; Text 'IW402'
   TextField "Text field_9" at 60,212 size 215x20; Text 'APT Confined Space Oxygen Level'
   TextField "Text field_10" at 7,212 size 53x20; Text 'IW404'
   TextField "Text field_13" at 60,250 size 215x20; Text 'RIO 7 Deck Main Pressure PT-415'
   TextField "Text field_14" at 7,250 size 53x20; Text 'IW408'
   TextField "Text field_15" at 60,288 size 215x20; Text 'APT BW Level LT-422-APT'
   TextField "Text field_16" at 7,288 size 53x20; Text 'IW410'
   TextField "Text field_26" at 928,114 size 62x18; Text 'Reading'
   TextField "Text field_27" at 1001,114 size 68x18; Text 'Low Low'
   TextField "Text field_28" at 1082,114 size 34x18; Text 'Low'
   TextField "Text field_29" at 1150,114 size 37x18; Text 'High'
   TextField "Text field_30" at 1203,114 size 74x18; Text 'High High'
   TextField "Text field_31" at 1076,92 size 74x18; Text 'Setpoints'
   TextField "Text field_65" at 702,138 size 215x20; Text 'APT BW ph TX-426-APT'
   IOField "I/O field_126" at 922,138 size 75x20; FormatPattern 99.9
      ProcessValue <- "20_TANKS_IP_DATA_RIO_07_FIRST_TANK_BWT_PH"
   TextField "Text field_66" at 649,138 size 53x20; Text 'IW416'
   TextField "Text field_67" at 702,175 size 215x20; Text 'APT BW Temperature 426-APT'
   IOField "I/O field_131" at 922,175 size 75x20; FormatPattern s999.9; Unit  °C
      ProcessValue <- "20_TANKS_IP_DATA_RIO_07_FIRST_TANK_BWT_TEMP"
   TextField "Text field_68" at 649,175 size 53x20; Text 'IW418'
   TextField "Text field_69" at 702,212 size 215x20; Text 'APT BW DO TX-428-APT'
   IOField "I/O field_136" at 922,212 size 75x20; FormatPattern s99.99; Unit  mg/l
      ProcessValue <- "20_TANKS_IP_DATA_RIO_07_FIRST_TANK_BWT_DO"
   TextField "Text field_70" at 649,212 size 53x20; Text 'IW420'
   TextField "Text field_71" at 702,249 size 215x20; Text 'RIO 7 Tanks Pressure PT-424'
   TextField "Text field_72" at 649,249 size 53x20; Text 'IW422'
   TextField "Text field_41" at 133,114 size 85x18; Text 'Description'
   TextField "Text field_42" at 771,114 size 85x18; Text 'Description'
   TextField "Text field_43" at 17,114 size 21x18; Text 'AI'
   TextField "Text field_44" at 661,114 size 21x18; Text 'AI'
   IOField "I/O field_21" at 281,250 size 75x20; FormatPattern 99.999; Unit  Bar
      ProcessValue <- "20_TANKS_IP_DATA_RIO_07_FIRST_TANK_DECK_IG_PRESS"
   IOField "I/O field_26" at 281,288 size 75x20; FormatPattern 999.9; Unit  %
      ProcessValue <- "20_TANKS_IP_DATA_RIO_07_FIRST_TANK_BWT_LEVEL"
   IOField "I/O field_93" at 922,249 size 75x20; FormatPattern s999.9; Unit  mBar
      ProcessValue <- "20_TANKS_IP_DATA_RIO_07_FIRST_TANK_TANKS_PRESS"
   IOField "I/O field_16" at 281,213 size 75x20; FormatPattern 99.9; Unit  %
      ProcessValue <- "20_TANKS_IP_DATA_RIO_07_FIRST_TANK_O2_MONITOR"
   IOField "I/O field_1" at 361,138 size 60x20; Authorization "User administration"; FormatPattern 999
      ProcessValue <- "2084_Setpoints_FIT418_LoLo"
   IOField "I/O field_3" at 429,138 size 60x20; Authorization "User administration"; FormatPattern 999
      ProcessValue <- "2084_Setpoints_FIT418_Lo"
   IOField "I/O field_4" at 497,138 size 60x20; Authorization "User administration"; FormatPattern 999
      ProcessValue <- "2084_Setpoints_FIT418_Hi"
   IOField "I/O field_5" at 565,138 size 60x20; Authorization "User administration"; FormatPattern 999
      ProcessValue <- "2084_Setpoints_FIT418_HiHi"
   IOField "I/O field_7" at 361,175 size 60x20; FormatPattern 999
      ProcessValue <- "2084_Setpoints_FIT420_LoLo"
   IOField "I/O field_8" at 429,175 size 60x20; FormatPattern 999
      ProcessValue <- "2084_Setpoints_FIT420_Lo"
   IOField "I/O field_9" at 497,175 size 60x20; Authorization "User administration"; FormatPattern 999
      ProcessValue <- "2084_Setpoints_FIT420_Hi"
   IOField "I/O field_10" at 565,175 size 60x20; Authorization "User administration"; FormatPattern 999
      ProcessValue <- "2084_Setpoints_FIT420_HiHi"
   IOField "I/O field_62" at 361,213 size 60x20; FormatPattern 99.9
      ProcessValue <- "2084_Setpoints_Conf O2 Level Lo Lo"
   IOField "I/O field_63" at 429,213 size 60x20; FormatPattern 99.9
      ProcessValue <- "2084_Setpoints_Conf O2 Level Lo"
   IOField "I/O field_64" at 496,213 size 60x20; Authorization "User administration"; FormatPattern 99.9
   IOField "I/O field_65" at 564,213 size 60x20; Authorization "User administration"; FormatPattern 99.9
   IOField "I/O field_22" at 361,250 size 60x20; FormatPattern 99.999
      ProcessValue <- "2084_Setpoints_PIT415_LoLo"
   IOField "I/O field_23" at 429,250 size 60x20; FormatPattern 99.999
      ProcessValue <- "2084_Setpoints_PIT415_Lo"
   IOField "I/O field_24" at 497,250 size 60x20; FormatPattern 99.999
      ProcessValue <- "2084_Setpoints_PIT415_Hi"
   IOField "I/O field_25" at 565,250 size 60x20; FormatPattern 99.999
      ProcessValue <- "2084_Setpoints_PIT415_HiHi"
   IOField "I/O field_30" at 429,287 size 60x20; Authorization "User administration"; FormatPattern 999
      ProcessValue <- "2084_Setpoints_LT422_Lo"
   IOField "I/O field_31" at 497,287 size 60x20; Authorization "User administration"; FormatPattern 999
      ProcessValue <- "2084_Setpoints_LT422_Hi"
   IOField "I/O field_32" at 361,287 size 60x20; FormatPattern 9.9
   IOField "I/O field_34" at 565,287 size 60x20; FormatPattern 9.9
   IOField "I/O field_52" at 1003,138 size 60x20; FormatPattern 99.9
   IOField "I/O field_53" at 1071,138 size 60x20; FormatPattern 99.9
      ProcessValue <- "2084_Setpoints_TX426 Port PH Lo"
   IOField "I/O field_54" at 1003,175 size 60x20; FormatPattern 99.9
   IOField "I/O field_55" at 1071,175 size 60x20; FormatPattern 99.9
   IOField "I/O field_57" at 1139,138 size 60x20; Authorization "User administration"; FormatPattern 99.9
      ProcessValue <- "2084_Setpoints_TX426 Port PH High"
   IOField "I/O field_58" at 1207,138 size 60x20; Authorization "User administration"; FormatPattern 99.9
   IOField "I/O field_59" at 1139,175 size 60x20; Authorization "User administration"; FormatPattern 99.9
   IOField "I/O field_60" at 1207,175 size 60x20; Authorization "User administration"; FormatPattern 99.9
   IOField "I/O field_89" at 1139,212 size 60x20; Authorization "User administration"; FormatPattern 99.9
      ProcessValue <- "2084_Setpoints_TX428 Port DO High"
   IOField "I/O field_90" at 1207,212 size 60x20; Authorization "User administration"; FormatPattern 99.9
   IOField "I/O field_91" at 1003,212 size 60x20; Authorization "User administration"; FormatPattern 99.9
   IOField "I/O field_92" at 1071,212 size 60x20; Authorization "User administration"; FormatPattern 99.9
      ProcessValue <- "2084_Setpoints_TX428 Port DO Lo"
   IOField "I/O field_94" at 1139,249 size 60x20; Authorization "User administration"; FormatPattern 999.9
      ProcessValue <- "2084_Setpoints_PIT424_Hi"
   IOField "I/O field_95" at 1207,249 size 60x20; Authorization "User administration"; FormatPattern 999.9
      ProcessValue <- "2084_Setpoints_PIT424_HiHi"
   IOField "I/O field_96" at 1004,249 size 60x20; Authorization "User administration"; FormatPattern 999.9
      ProcessValue <- "2084_Setpoints_PIT424_LoLo"
   IOField "I/O field_97" at 1072,249 size 60x20; Authorization "User administration"; FormatPattern 999.9
      ProcessValue <- "2084_Setpoints_PIT424_Lo"
   Group "Group" at 455,41 size 373x50
   Button "HmiScreenItemData_8" at 469,45 size 355x40; TextOn 'Back'; TextOff 'Text'
   TextField "Screen title" at 455,41 size 373x50; Text 'Screen title'

